(* Logix 5000 project; controller OWF Emulate 5570 rev 30.12; software revision 30.00; part 4 of 4 *)
(* MainProgram, continued *)

ROUTINE OWF_Test   (* structured text *)
   
   
   Jsr(Original_OWF);
   
   
   
   
END_ROUTINE
END_PROGRAM
